// TIA Portal project "KO_CHLab2" (V13)

(* hardware
DEVICE "S7-1200 station_1"  S7-1200 Station
   slot 0: "Rack_0"  Rack  V1.0
   slot 1: "PLC_1"  CPU 1214C AC/DC/Rly  6ES7 214-1BE30-0XB0  V2.2
*)

// ===== PLC "PLC_1"  CPU 1214C AC/DC/Rly =====

VAR_GLOBAL   // PLC tag table "Default tag table"
   "Clock_Byte" AT %MB0 : Byte;
   "Clock_10Hz" AT %M0.0 : Bool;
   "Clock_5Hz" AT %M0.1 : Bool;
   "Clock_2.5Hz" AT %M0.2 : Bool;
   "Clock_2Hz" AT %M0.3 : Bool;
   "Clock_1.25Hz" AT %M0.4 : Bool;
   "Clock_1Hz" AT %M0.5 : Bool;
   "Clock_0.625Hz" AT %M0.6 : Bool;
   "Clock_0.5Hz" AT %M0.7 : Bool;
   "ret_val" AT %MW2 : Int;
   "Tag_1" AT %I0.0 : Bool;
   "Tag_2" AT %M10.1 : Bool;
END_VAR

DATA_BLOCK "Danelogowania"   // DB3
{ S7_Optimized_Access := 'FALSE' }
VERSION : 0.1
   VAR
      Admin : Struct
      END_STRUCT;
      spr_admin : Bool;
      spr_user : Bool;
      log : String;
      i : Int;
      has : String;
      spr : Bool;
      Users : Array[0..11] of Struct
      END_STRUCT;
      Umowy : Array[0..11] of Struct
      END_STRUCT;
      tankowane_paliwo : Int;
      podlaczone : Bool;
      starttank : Bool;
      stoptank : Bool;
      indeksu : Int;
      user_nr : Int;
      limit : Int;
      userhas : String;
      userlog : String;
      userpaliwo : Int;
      startnocny : Bool;
      myint : Int;
   END_VAR
BEGIN
END_DATA_BLOCK

// folder: System blocks/Program resources

DATA_BLOCK "IEC_Counter_0_DB"   // DB1
{ S7_Optimized_Access := 'FALSE' }
AUTHOR : Simatic
FAMILY : IEC
NAME : CNTR
VERSION : 1.0
// stored: InstanceOfName ?
"?"
BEGIN
END_DATA_BLOCK

// folder: (top level)

ORGANIZATION_BLOCK "Main"   // OB1, LAD, ProgramCycle
TITLE = "Main Program Sweep (Cycle)"
{ S7_Optimized_Access := 'FALSE' }
VERSION : 0.1
   VAR_TEMP   // added for the SCL form of the ladder/FBD networks
      _w1 : Bool;
      _w2 : Bool;
   END_VAR
BEGIN

REGION Network 1
   // Polaczenie z web serwerwem naszej strony
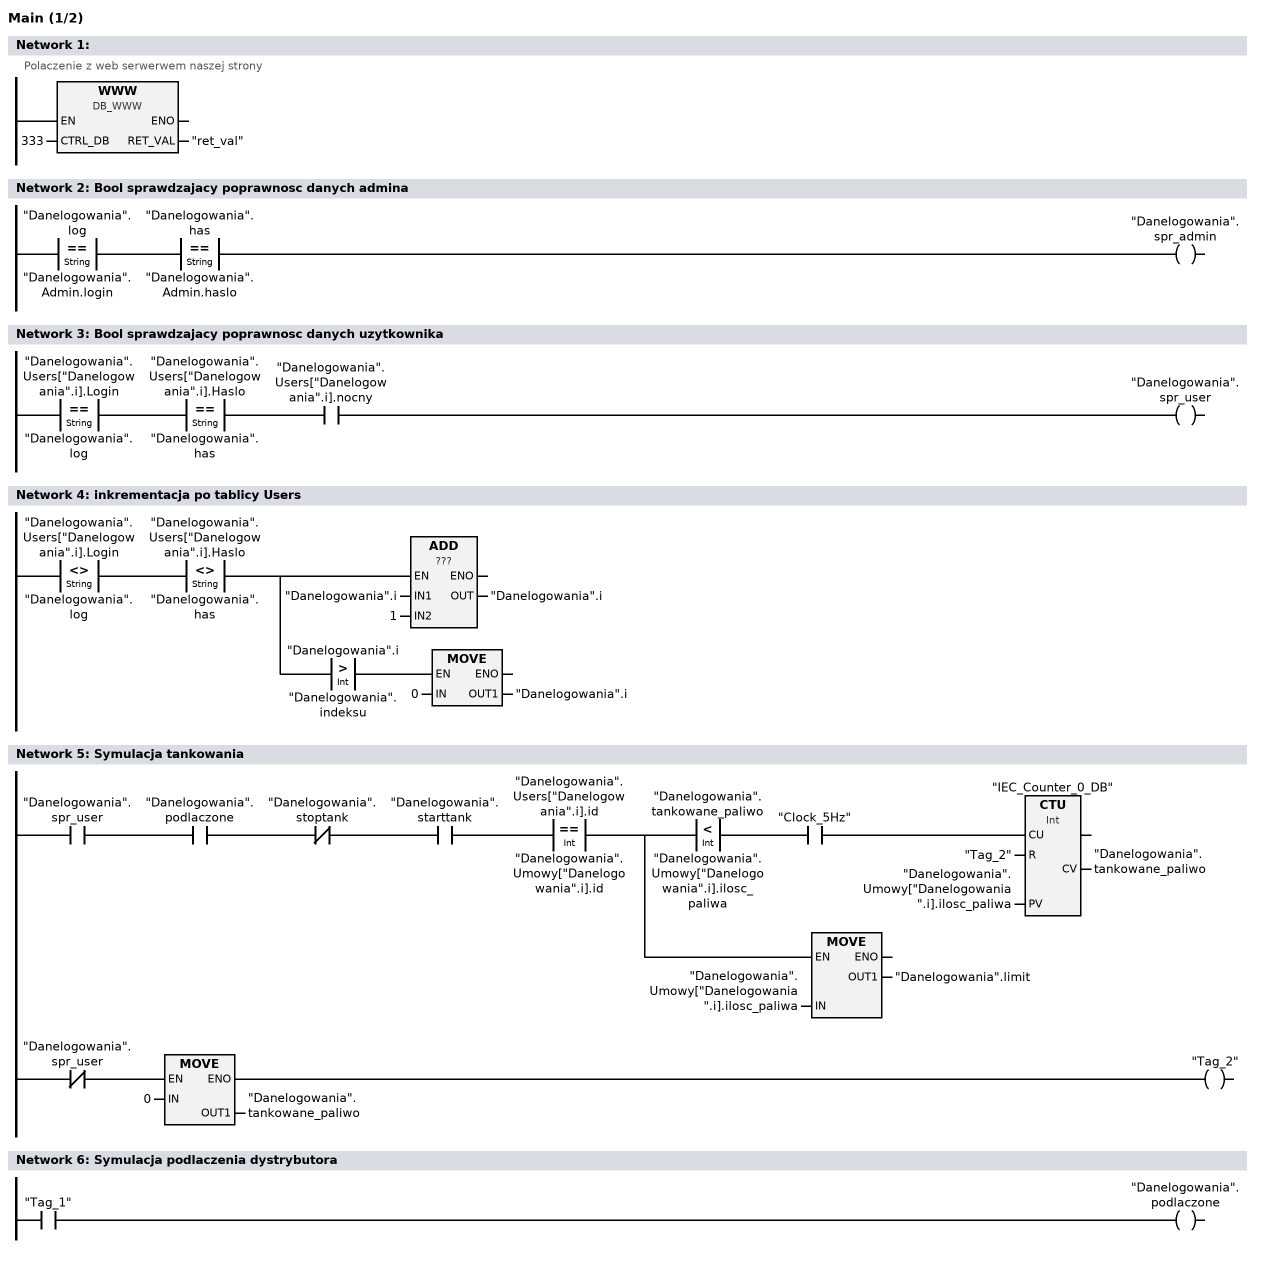
   "ret_val" := WWW(CTRL_DB := 333);
END_REGION

REGION Network 2: Bool sprawdzajacy poprawnosc danych admina
   RUNG wire#powerrail
      { S7_Templates := "SrcType := String" } EQ_Contact(in1 := "Danelogowania".log, in2 := "Danelogowania".Admin.login)
      { S7_Templates := "SrcType := String" } EQ_Contact(in1 := "Danelogowania".has, in2 := "Danelogowania".Admin.haslo)
      Coil( "Danelogowania".spr_admin )
   END_RUNG
   // the same network as SCL:
   "Danelogowania".spr_admin := ("Danelogowania".log = "Danelogowania".Admin.login) AND ("Danelogowania".has = "Danelogowania".Admin.haslo);
END_REGION

REGION Network 3: Bool sprawdzajacy poprawnosc danych uzytkownika
   RUNG wire#powerrail
      { S7_Templates := "SrcType := String" } EQ_Contact(in1 := "Danelogowania".Users["Danelogowania".i].Login, in2 := "Danelogowania".log)
      { S7_Templates := "SrcType := String" } EQ_Contact(in1 := "Danelogowania".Users["Danelogowania".i].Haslo, in2 := "Danelogowania".has)
      Contact( "Danelogowania".Users["Danelogowania".i].nocny )
      Coil( "Danelogowania".spr_user )
   END_RUNG
   // the same network as SCL:
   "Danelogowania".spr_user := ("Danelogowania".Users["Danelogowania".i].Login = "Danelogowania".log) AND ("Danelogowania".Users["Danelogowania".i].Haslo = "Danelogowania".has) AND "Danelogowania".Users["Danelogowania".i].nocny;
END_REGION

REGION Network 4: inkrementacja po tablicy Users
   RUNG wire#powerrail
      { S7_Templates := "SrcType := String" } NE_Contact(in1 := "Danelogowania".Users["Danelogowania".i].Login, in2 := "Danelogowania".log)
      { S7_Templates := "SrcType := String" } NE_Contact(in1 := "Danelogowania".Users["Danelogowania".i].Haslo, in2 := "Danelogowania".has)
      wire#w1
      { S7_Templates := "SrcType := ???"; S7_GenerateENO := "TRUE" } Add(in1 := "Danelogowania".i, in2 := 1, out => "Danelogowania".i)
   END_RUNG
   RUNG wire#w1
      { S7_Templates := "SrcType := Int" } GT_Contact(in1 := "Danelogowania".i, in2 := "Danelogowania".indeksu)
      { S7_GenerateENO := "TRUE" } Move(in := 0, out1 => "Danelogowania".i)
   END_RUNG
   // the same network as SCL:
   #_w1 := ("Danelogowania".Users["Danelogowania".i].Login <> "Danelogowania".log) AND ("Danelogowania".Users["Danelogowania".i].Haslo <> "Danelogowania".has);
   IF #_w1 THEN "Danelogowania".i := "Danelogowania".i + 1; END_IF;
   IF #_w1 AND ("Danelogowania".i > "Danelogowania".indeksu) THEN "Danelogowania".i := 0; END_IF;
END_REGION

REGION Network 5: Symulacja tankowania
   // ENO of a box is taken as its EN; it also drops when the box reports an error
   #_w1 := "Danelogowania".spr_user AND "Danelogowania".podlaczone AND NOT "Danelogowania".stoptank AND "Danelogowania".starttank AND ("Danelogowania".Users["Danelogowania".i].id = "Danelogowania".Umowy["Danelogowania".i].id);
   "IEC_Counter_0_DB".CTU(CU := #_w1 AND ("Danelogowania".tankowane_paliwo < "Danelogowania".Umowy["Danelogowania".i].ilosc_paliwa) AND "Clock_5Hz",
                          R := "Tag_2",
                          PV := "Danelogowania".Umowy["Danelogowania".i].ilosc_paliwa,
                          CV => "Danelogowania".tankowane_paliwo);
   IF #_w1 THEN "Danelogowania".limit := "Danelogowania".Umowy["Danelogowania".i].ilosc_paliwa; END_IF;
   #_w2 := NOT "Danelogowania".spr_user;
   IF #_w2 THEN "Danelogowania".tankowane_paliwo := 0; END_IF;
   "Tag_2" := #_w2;
END_REGION

REGION Network 6: Symulacja podlaczenia dystrybutora
   RUNG wire#powerrail
      Contact( "Tag_1" )
      Coil( "Danelogowania".podlaczone )
   END_RUNG
   // the same network as SCL:
   "Danelogowania".podlaczone := "Tag_1";
END_REGION

REGION Network 7: Przypisywanie do rozpiski nocnych
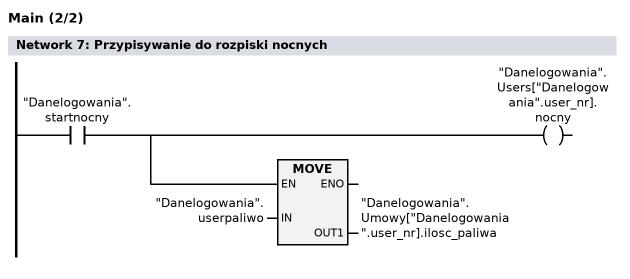
   RUNG wire#powerrail
      Contact( "Danelogowania".startnocny )
      wire#w1
      Coil( "Danelogowania".Users["Danelogowania".user_nr].nocny )
   END_RUNG
   RUNG wire#w1
      { S7_GenerateENO := "TRUE" } Move(in := "Danelogowania".userpaliwo, out1 => "Danelogowania".Umowy["Danelogowania".user_nr].ilosc_paliwa)
   END_RUNG
   // the same network as SCL:
   "Danelogowania".Users["Danelogowania".user_nr].nocny := "Danelogowania".startnocny;
   IF "Danelogowania".startnocny THEN
       "Danelogowania".Umowy["Danelogowania".user_nr].ilosc_paliwa := "Danelogowania".userpaliwo;
   END_IF;
END_REGION
END_ORGANIZATION_BLOCK